screen "SettingPrinter" 800x414, template "Template_Mirai"
   on GenerateScreen: SetTag("screen_titles", 52)
   Button "Button_3" at 256,226 size 80x40; TextOff 'Connect / Pripoj'
      on Release: ResetBit("CON_ConnectHMI")
      on Press: SetBit("CON_ConnectHMI")
   TextField "Text field_3" at 19,231 size 25x32; Text 'IP'
   IOField "I/O field_1" at 61,231 size 180x32; FormatPattern ????????????????????
      ProcessValue <- "PrinterData_CON_PrinterBagData_RemoteAddress"
   TextField "Text field_4" at 167,152 size 42x32; Text 'CON'
   SymbolicIOField "Symbolic I/O field_1" at 65,186 size 170x32; TextOn '1'; TextOff '0'; TextList "CON_Printers"
      ProcessValue <- "PrinterData_CON_PrinterSelection"
   Button "Button_6" at 256,42 size 80x40; TextOff 'Connect / Pripoj'
      on Release: ResetBit("TRP_ConnectHMI")
      on Press: SetBit("TRP_ConnectHMI")
   Button "Button_1" at 256,98 size 120x40; TextOff 'Initialization / Inicializácia'
      on Release: ResetBit("PrinterData_TRP_PrinterData_Initialization")
      on Press: SetBit("PrinterData_TRP_PrinterData_Initialization")
   TextField "Text field_1" at 168,8 size 42x32; Text 'TRP'
   TextField "Text field_2" at 13,47 size 25x32; Text 'IP'
   IOField "I/O field_5" at 38,47 size 213x32; FormatPattern ????????????????????
      ProcessValue <- "PrinterData_TRP_PrinterData_RemoteAddress"
   IOField "I/O field_2" at 61,303 size 180x32; FormatPattern ????????????????????????????????????????????????????????????????????????????????
      ProcessValue <- "PrinterData_CON_PrinterBagData_NonMDR_LabelName"
   TextField "Text field_5" at 19,274 size 223x32; Text 'Non-MDR label name'
   Button "Button_5" at 672,302 size 120x40; TextOff 'Camera settings Nastavenia kamery'
      on Release: ActivateScreen("Setting_DelayTimeM", 0)
   GraphicView "Graphic view_1" at 348,42 size 44x30; Picture "Wbox"
      Visibility <- "TRP_DB_MarkemImaje_ConnectionStatus"
   GraphicView "Graphic view_2" at 346,43 size 45x27; Picture "Cbox"
      Visibility <- "TRP_DB_MarkemImaje_ConnectionStatus"
   GraphicView "Graphic view_3" at 348,229 size 44x30; Picture "Wbox"
      Visibility <- "CON_PrinterConnection"
   GraphicView "Graphic view_4" at 347,231 size 45x27; Picture "Cbox"
      Visibility <- "CON_PrinterConnection"
   Button "Button_4" at 257,301 size 120x40; TextOff 'Initialization / Inicializácia'
      on Release: ResetBit("PrinterData_CON_PrinterBagData_Initialization")
      on Press: SetBit("PrinterData_CON_PrinterBagData_Initialization")
   Switch "Switch_1" at 115,82 size 120x56; TextOn 'DOLE'; CaptionText 'Inverse / Obratena tlac'; TextOff 'HORE'
      on SwitchOff: ResetBit("PrinterData_TRP_PrinterData_Inverse")
      on SwitchOn: SetBit("PrinterData_TRP_PrinterData_Inverse")
      ProcessValue <- "PrinterData_TRP_PrinterData_Inverse"

screen "Setting_DelayTimeM" 800x414, template "Template_Mirai"
   on GenerateScreen: SetTag("screen_titles", 53)
   IOField "I/O field_2" at 160,63 size 104x40; FormatPattern 999
      ProcessValue <- "SP_HMI_Box_Cam_Delay_time_trigger"
   TextField "Text field_2" at 4,63 size 148x40; Text '2D Code Box / 2D kód krabice'
   TextField "Text field_3" at 160,16 size 104x40; Text 'Trigger delay (ms) Oneskorenie čítania (ms)'
   Button "Btn_OpenEditor" at 4,313 size 160x32; TextOff 'Back / Späť'
      on Click: ActivateScreen("SettingPrinter", 0)
   Button "Btn_OpenEditor_1" at 180,313 size 160x32; TextOff 'Camera position / Pozícia kamery'; Authorization "Operate"
      on Click: ActivateScreen("Setting_CameraM", 0)

screen "StatusM" 800x414, template "Template_Mirai"
   on GenerateScreen: SetTag("screen_titles", 51)
   TextField "Text field_2" at 28,39 size 43x23; Text '(01)'
   TextField "Text field_3" at 28,77 size 43x23; Text '(10)'
   TextField "Text field_4" at 28,115 size 43x23; Text '(91)'
   TextField "Text field_5" at 28,153 size 43x23; Text '(92)'
   TextField "Text field_6" at 28,191 size 43x23; Text '(11)'
   TextField "Text field_7" at 28,229 size 43x23; Text '(15)'
   IOField "I/O field_1" at 81,33 size 171x34; FormatPattern ????????????????????????????????????????????????????????????????????????????????
      ProcessValue <- "OPC_TRP_Materia_ActualGTIN_Number"
   IOField "I/O field_2" at 81,71 size 171x34; FormatPattern ????????????????????????????????????????????????????????????????????????????????
      ProcessValue <- "OPC_TRP_Materia_ActualBatchNumber"
   TextField "Text field_8" at 171,9 size 42x23; Text 'TRP'
   IOField "I/O field_3" at 81,109 size 171x34; FormatPattern ????????????????????????????????????????????????????????????????????????????????
      ProcessValue <- "OPC_TRP_Materia_ActualAricleNumber"
   IOField "I/O field_4" at 81,147 size 171x34; FormatPattern ??????
      ProcessValue <- "PrinterData_CON_PrinterBagData_Time"
   IOField "I/O field_5" at 81,185 size 171x34; FormatPattern ????????????????????????????????????????????????????????????????????????????????
      ProcessValue <- "PrinterData_CON_PrinterBagData_Date"
   IOField "I/O field_6" at 81,223 size 171x34; FormatPattern ??????????
      ProcessValue <- "TRP_DB_MarkemImaje_ExtDate"
   TextField "Text field_1" at 548,10 size 110x23; Text 'PLAIN Data'
   TextField "Text field_11" at 400,33 size 90x23; Text 'EAN_TRP / EAN TRP'
   TextField "Text field_13" at 400,63 size 56x23; Text 'Batch'
   TextField "Text field_15" at 400,93 size 100x23; Text 'MachineID'
   TextField "Text field_16" at 400,123 size 90x23; Text 'MDR Flag'
   TextField "Text field_17" at 400,153 size 66x23; Text 'Article'
   TextField "Text field_18" at 400,183 size 99x23; Text 'Batch END'
   TextField "Text field_19" at 400,214 size 92x23; Text 'ART Base'
   TextField "Text field_20" at 400,246 size 87x23; Text 'ART Flag'
   TextField "Text field_21" at 400,278 size 110x23; Text 'Market Reg'
   TextField "Text field_22" at 400,310 size 42x23; Text 'BBD'
   IOField "I/O field_11" at 570,32 size 200x25; FormatPattern ??????????????
      ProcessValue <- "OPC_TRP_Materia_NewGTIN_Number"
   IOField "I/O field_12" at 570,62 size 200x25; FormatPattern ????????????????????????????????????????????????????????????????????????????????
      ProcessValue <- "OPC_CON_Material_NewBatchNumber"
   IOField "I/O field_13" at 570,92 size 200x25; FormatPattern ????????????????????????????????????????????????????????????????????????????????
      ProcessValue <- "OPC_TRP_Materia_NewMachineID"
   IOField "I/O field_14" at 570,122 size 200x25; FormatPattern ????????????????????????????????????????????????????????????????????????????????
      ProcessValue <- "OPC_CON_Material_NewMDR_Flag"
   IOField "I/O field_15" at 570,152 size 200x25; FormatPattern 9999999999
      ProcessValue <- "OPC_TRP_Materia_NewArticleNumber"
   IOField "I/O field_16" at 570,182 size 200x25; FormatPattern ????????????????????????????????????????????????????????????????????????????????
      ProcessValue <- "OPC_CON_Material_NewBatchEndTime"
   IOField "I/O field_17" at 570,213 size 200x25; FormatPattern 9999999999
      ProcessValue <- "OPC_CON_Material_NewArtBaseNumber"
   IOField "I/O field_18" at 570,245 size 200x25; FormatPattern ????????????????????????????????????????????????????????????????????????????????
      ProcessValue <- "OPC_CON_Material_NewArticleFlag"
   IOField "I/O field_19" at 570,277 size 200x25; FormatPattern ?????????????????????
      ProcessValue <- "OPC_CON_Material_NewMarketREG_Code"
   IOField "I/O field_20" at 570,309 size 200x25; FormatPattern ????????????????????????????????????????????????????????????????????????????????
      ProcessValue <- "OPC_CON_Material_NewBBD"
   IOField "I/O field_7" at 55,284 size 115x32; HelpText 'Enter ip+port 10.176.48.110:45'; FormatPattern ??????????
      ProcessValue <- "OPC_TRP_Materia_ActualBatchNumber"
   IOField "I/O field_8" at 194,284 size 115x32; HelpText 'Enter ip+port 10.176.48.110:45'; FormatPattern ??????????
      ProcessValue <- "OPC_CON_Material_ActualArtBaseNumber"
      Visibility <- "CON_DB_HandleComBag_ActualArtFlag"
   IOField "I/O field_10" at 20,302 size 115x32; HelpText 'Enter ip+port 10.176.48.110:45'; FormatPattern ??????????
      ProcessValue <- "OPC_CON_Material_ActualMarketRegCode"
   TextField "Text field_14" at 127,307 size 42x23; Text 'BBD'
      Visibility <- "TRP_DB_MarkemImaje_ExpFlag"
   IOField "I/O field_9" at 165,303 size 76x32; HelpText 'Enter ip+port 10.176.48.110:45'; FormatPattern ??????
      ProcessValue <- "OPC_CON_Material_ActualBBD"
   IOField "I/O field_23" at 296,284 size 76x32; HelpText 'Enter ip+port 10.176.48.110:45'; FormatPattern ?????
      ProcessValue <- "TRP_DB_MarkemImaje_TimePrinted"
      Visibility <- "CON_DB_HandleComBag_ActualArtFlag"
   IOField "I/O field_24" at 159,284 size 76x32; HelpText 'Enter ip+port 10.176.48.110:45'; FormatPattern ??????
      ProcessValue <- "TRP_DB_MarkemImaje_TimePrinted"
      Visibility <- "CON_DB_HandleComBag_ActualArtFlag"
   TextField "Text field_9" at 20,288 size 40x23; Text 'LOT'
   TextField "Text field_12" at 159,288 size 43x23; Text 'ART'
      Visibility <- "CON_DB_HandleComBag_ActualArtFlag"
   TextField "Text field_10" at 151,263 size 43x23; Text 'CON'
   IOField "I/O field_21" at 150,152 size 44x23; HelpText 'Enter ip+port 10.176.48.110:45'; FormatPattern ???
      ProcessValue <- "OPC_TRP_Materia_ActualMachineID"
   IOField "I/O field_22" at 188,152 size 58x23; HelpText 'Enter ip+port 10.176.48.110:45'; FormatPattern 99999
      ProcessValue <- "TRP_DB_MarkemImaje_Serial"

screen "Rec_Edit" 800x414, template "Template_Enigma"
   on GenerateScreen: SetTag("screen_titles", 6)
   IOField "I/O field_1" at 407,54 size 104x32; Authorization "Recipe management"; FormatPattern 9999
      ProcessValue <- "Rec_HMI_Bag_Cam_Vertiacal_position"
   IOField "I/O field_2" at 407,131 size 104x32; Authorization "Recipe management"; FormatPattern s999
      ProcessValue <- "Rec_HMI_Bag_Cam_Angle"
   IOField "I/O field_3" at 407,93 size 104x32; Authorization "Recipe management"; FormatPattern 9999
      ProcessValue <- "Rec_HMI_Bag_Cam_Horizontal_position"
   TextField "Text field_1" at 299,54 size 104x32; Text 'A'
   TextField "Text field_2" at 299,93 size 104x32; Text 'B'
   TextField "Text field_3" at 299,131 size 104x32; Text 'C'
   TextField "Text field_4" at 623,54 size 36x32; Text 'mm'
   TextField "Text field_5" at 623,93 size 36x32; Text 'mm'
   TextField "Text field_6" at 623,131 size 36x32; Text '°'
   TextField "Text field_15" at 299,167 size 104x40; Text 'Trigger delay Oneskorenie čítania'
   IOField "I/O field_4" at 407,171 size 104x32; Authorization "Recipe management"; FormatPattern 999
      ProcessValue <- "Rec_HMI_Bag_Cam_Delay_time_trigger"
   IOField "I/O field_5" at 515,171 size 104x32; Authorization "Recipe management"; FormatPattern 999
      ProcessValue <- "Rec_HMI_Box_Cam_Delay_time_trigger"
   TextField "Text field_16" at 623,171 size 36x32; Text 'ms'
   TextField "Text field_18" at 419,18 size 80x32; Text 'BAG / SÁČOK'
   TextField "Text field_19" at 527,18 size 80x32; Text 'BOX / KRABICA'
   IOField "I/O field_8" at 515,54 size 104x32; Authorization "Recipe management"; FormatPattern 9999
      ProcessValue <- "Rec_HMI_Box_Cam_Vertiacal_position"
   IOField "I/O field_9" at 515,131 size 104x32; Authorization "Recipe management"; FormatPattern s999
      ProcessValue <- "Rec_HMI_Box_Cam_Angle"
   IOField "I/O field_10" at 515,93 size 104x32; Authorization "Recipe management"; FormatPattern 9999
      ProcessValue <- "Rec_HMI_Box_Cam_Horizontal_position"
   Button "Btn_Save" at 692,8 size 80x32; TextOff 'SAVE / ULOŽ'; Authorization "Recipe management"
      on Click: SetTag("Rec_FunctionUsed", 7); "Rec_SafeSave"()
   Button "Btn_ExitEditor" at 8,313 size 216x32; TextOff 'Exit recipe editor / Ukonči editor receptov'
      on Click: ActivateScreen("Rec_Overview", 0)
   GraphicView "Graphic view_1" at 20,77 size 222x229; Picture "CognexDatamanClearedAndSemiTransparent2"
   TextField "Text field_10" at 18,184 size 32x40; Text 'A'
   TextField "Text field_11" at 102,71 size 32x40; Text 'B'
   TextField "Text field_12" at 179,78 size 32x40; Text 'C'
   Button "Btn_ReadSP" at 668,72 size 124x32; TextOff 'READ from PLC / NAČÍTAJ z PLC'; Authorization "Recipe management"
      on Click: SetTag("Rec_FunctionUsed", 8); function_b456aad1(1, "Rec_ReadSPResult")
   TextField "Text field_7" at 8,8 size 264x62; Text 'Recipe name: / Názov receptu: / 配方名'
   IOField "I/O field_6" at 14,35 size 252x30; Authorization "Recipe management"; FormatPattern ????????????????????????????????????????
      ProcessValue <- "Rec_SelectedRecipe"
   GraphicIOField "Graphic I/O field_1" at 408,250 size 32x32; PictureList "On_Off_Editable"
      ProcessValue <- "Rec_HMI_Enigma_off"
   Button "Button_1" at 408,250 size 32x32; TextOff 'Text'
      on Click: InvertBit("Rec_HMI_Enigma_off")
   IOField "I/O field_7" at 407,211 size 104x32; Authorization "Recipe management"; FormatPattern 9999
      ProcessValue <- "Rec_HMI_Bag_Cam_Fps"
   TextField "Text field_13" at 299,211 size 104x32; Text 'Num of pics / Počet snímok'
   IOField "I/O field_11" at 515,211 size 104x32; Authorization "Recipe management"; FormatPattern 9999
      ProcessValue <- "Rec_HMI_Box_Cam_Fps"
   TextField "Text field_14" at 299,250 size 104x32; Text 'Enigma'
   GraphicIOField "Graphic I/O field_2" at 624,250 size 32x32; PictureList "On_Off_Editable"
      ProcessValue <- "Rec_HMI_Mirai_off"
   Button "Button_2" at 624,250 size 32x32; TextOff 'Text'
      on Click: InvertBit("Rec_HMI_Mirai_off")
   TextField "Text field_20" at 515,250 size 104x32; Text 'Mirai'
   Button "Btn_OK_Save_NoNameSpecified" at 692,313 size 80x32; TextOff 'OK / 确定'
      on Click: SetTag("Rec_SaveResult", 0)
      Visibility <- "Rec_SaveResult"
   TextField "Text field_17" at 288,292 size 376x53; Text 'No recipe name set, recipe not saved. Set recipe name and try again. Žiaden zadaný názov receptu, recept sa neuložil. Nastavte názov receptu a skúste to znova. 未设置配方名 不能保存配方。 输入配方名再保存。'
      Visibility <- "Rec_SaveResult"
   TextField "Text field_8" at 288,292 size 376x53; Text 'Saving recipe ... / Ukladanie receptu ... / 配方保存中…'
      Visibility <- "Rec_SaveResult"
   Button "Btn_OK_Save_Success" at 692,313 size 80x32; TextOff 'OK / 确定'
      on Click: SetTag("Rec_SaveResult", 0)
      Visibility <- "Rec_SaveResult"
   TextField "Text field_9" at 288,292 size 376x53; Text 'Recipe saving succeeded. Ukladanie receptu bolo úspešné. 保存配方 成功。'
      Visibility <- "Rec_SaveResult"
   TextField "Text field_24" at 288,292 size 376x53; Text 'Recipe saving failed. Ukladanie receptu zlyhalo. 保存配方 失败。'
      Visibility <- "Rec_SaveResult"
   Button "Btn_OK_Save_Fail" at 692,313 size 80x32; TextOff 'OK / 确定'
      on Click: SetTag("Rec_SaveResult", 0)
      Visibility <- "Rec_SaveResult"
   TextField "Text field_25" at 288,292 size 376x53; Text 'Reading setpoints ... / Čítanie požadovaných hodnôt ... / 读取设定值…'
      Visibility <- "Rec_ReadSPResult"
   Button "Btn_OK_ReadSP_Success" at 692,313 size 80x32; TextOff 'OK / 确定'
      on Click: SetTag("Rec_ReadSPResult", 0)
      Visibility <- "Rec_ReadSPResult"
   TextField "Text field_26" at 288,292 size 376x53; Text 'Reading of setpoints succeeded. Čítanie požadovaných hodnôt bolo úspešné. 读取设定值 成功。'
      Visibility <- "Rec_ReadSPResult"
   TextField "Text field_27" at 288,292 size 376x53; Text 'Reading of setpoints failed. Čítanie požadovaných hodnôt zlyhalo. 读取设定值 失败。'
      Visibility <- "Rec_ReadSPResult"
   Button "Btn_OK_ReadSP_Fail" at 692,313 size 80x32; TextOff 'OK / 确定'
      on Click: SetTag("Rec_ReadSPResult", 0)
      Visibility <- "Rec_ReadSPResult"
   Rectangle "Rectangle_2" at 0,0 size 800x414
      Visibility <- "Rec_FunctionResultSwitch"

screen "Rec_Overview" 800x414, template "Template_Enigma"
   on GenerateScreen: SetTag("screen_titles", 4); SetTag("Rec_FunctionUsed", 0)
   RecipeView "Recipe view_1" at 4,44 size 792x80; DataRecordNameCaption 'Select recipe: / Vyber recept:'; Tag4DataRecord "Rec_SelectedRecipe"; Recipe "ReaderRecipes"
      Visibility <- "Rec_FunctionResultSwitch"
   Button "Btn_Edit" at 88,136 size 76x32; TextOff 'EDIT UPRAV 编辑 所选 配方'; Authorization "Recipe management"
      on Click: SetTag("Rec_FunctionUsed", 5); "Rec_SafeEdit"()
   Button "Btn_Load" at 636,136 size 160x32; TextOff 'LOAD to PLC NAHRAJ do PLC 下载 所选 配方 到PLC'; Authorization "Operate"
      on Click: SetTag("Rec_FunctionUsed", 1); "Rec_SafeLoad"()
   Button "Btn_Delete" at 362,136 size 76x32; TextOff 'DELETE VYMAŽ 删除 所选 配方'; Authorization "Recipe management"
      on Click: SetTag("Rec_FunctionUsed", 2); "Rec_SafeDelete"()
   Button "Btn_View" at 4,136 size 76x32; TextOff 'VIEW ZOBRAZ 浏览 所选 配方'; Authorization "Operate"
      on Click: SetTag("Rec_FunctionUsed", 6); "Rec_SafeView"()
   Button "Btn_OpenEditor" at 4,313 size 216x32; TextOff 'Open recipe editor / Otvor editor receptov'; Authorization "Recipe management"
      on Click: SetTag("Rec_SelectedRecipe", ''); ActivateScreen("Rec_Edit", 0)
   TextField "Text field_12" at 8,8 size 201x32; Text 'Article number: / Číslo artiklu:'
   IOField "I/O field_6" at 200,8 size 162x32; FormatPattern ??????????
      ProcessValue <- "PlainHandle_DB_NewArticleNum"
   Button "Btn_OK_Edit_NoRecipeSelected" at 362,176 size 76x32; TextOff 'OK / 确定'
      on Click: SetTag("Rec_EditResult", 0)
      Visibility <- "Rec_EditResult"
   Button "Btn_OK_Delete_NoRecipeSelected" at 362,176 size 76x32; TextOff 'OK / 确定'
      on Click: SetTag("Rec_DeleteResult", 0)
      Visibility <- "Rec_DeleteResult"
   Button "Btn_OK_View_NoRecipeSelected" at 362,176 size 76x32; TextOff 'OK / 确定'
      on Click: SetTag("Rec_ViewResult", 0)
      Visibility <- "Rec_ViewResult"
   Button "Btn_OK_Load_NoRecipeSelected" at 362,176 size 76x32; TextOff 'OK / 确定'
      on Click: SetTag("Rec_LoadResult", 0)
      Visibility <- "Rec_LoadResult"
   TextField "Text field_15" at 4,44 size 792x124; Text 'No recipe selected. / Nie je vybratý žiaden recept. / 未选配方。'
      Visibility <- "Rec_FunctionResultSwitch"
   TextField "Text field_11" at 4,44 size 792x124; Text 'Recipe loading failed. / Načítavanie receptu zlyhalo. / 下载配方失败。'
      Visibility <- "Rec_LoadResult"
   Button "Btn_OK_Load_Fail" at 362,176 size 76x32; TextOff 'OK / 确定'
      on Click: SetTag("Rec_LoadResult", 0)
      Visibility <- "Rec_LoadResult"
   TextField "Text field_7" at 4,44 size 792x124; Text 'Recipe deletion failed. / Mazanie receptu zlyhalo. / 删除配方失败。'
      Visibility <- "Rec_DeleteResult"
   Button "Btn_OK_Delete_Fail" at 362,176 size 76x32; TextOff 'OK / 确定'
      on Click: SetTag("Rec_DeleteResult", 0)
      Visibility <- "Rec_DeleteResult"
   Rectangle "Rectangle_1" at 0,0 size 800x414
      Visibility <- "Rec_FunctionResultSwitch"
   TextField "Text field_4" at 4,44 size 792x124; Text 'Recipe loading ... / Načítavanie receptu... / 配方表下载中…'
      Visibility <- "Rec_LoadResult"
   Button "Btn_OK_Load_Success" at 362,176 size 76x32; TextOff 'OK / 确定'
      on Click: SetBit("HMI_Control_NewRecipeLoaded"); SetTag("Rec_LoadResult", 0)
      Visibility <- "Rec_LoadResult"
   TextField "Text field_3" at 4,44 size 792x124; Text 'Recipe loading succeeded. / Načítavanie receptu bolo úspešné. / 下载配方成功。'
      Visibility <- "Rec_LoadResult"
   TextField "Text field_5" at 4,44 size 792x124; Text 'Deleting recipe ... / Vymazávanie receptu... / 删除配方…'
      Visibility <- "Rec_DeleteResult"
   Button "Btn_OK_Delete_Success" at 362,176 size 76x32; TextOff 'OK / 确定'
      on Click: SetTag("Rec_SelectedRecipe", ''); SetTag("Rec_DeleteResult", 0)
      Visibility <- "Rec_DeleteResult"
   TextField "Text field_6" at 4,44 size 792x124; Text 'Recipe deletion succeeded. / Mazanie receptu bolo úspešné. / 删除配方成功。'
      Visibility <- "Rec_DeleteResult"
   TextField "Text field_16" at 4,44 size 792x124; Text 'Opening recipe for editing ... / Prebieha otváranie receptu na úpravu ... / 打开编辑配方…'
      Visibility <- "Rec_EditResult"
   Button "Btn_OK_Edit_Success" at 362,176 size 76x32; TextOff 'OK / 确定'
      on Click: SetTag("Rec_EditResult", 0); ActivateScreen("Rec_Edit", 2)
      Visibility <- "Rec_EditResult"
   TextField "Text field_17" at 4,44 size 792x124; Text 'Recipe opening for editing succeeded. / Otváranie receptu na úpravu bolo úspešné. / 打开编辑配方成功。'
      Visibility <- "Rec_EditResult"
   TextField "Text field_1" at 4,44 size 792x124; Text 'Recipe opening for editing failed. / Otváranie receptu na úpravu zlyhalo. / 打开编辑配方失败。'
      Visibility <- "Rec_EditResult"
   Button "Btn_OK_Edit_Fail" at 362,176 size 76x32; TextOff 'OK / 确定'
      on Click: SetTag("Rec_EditResult", 0)
      Visibility <- "Rec_EditResult"
   TextField "Text field_2" at 4,44 size 792x124; Text 'Opening recipe for viewing ... / Prebieha otváranie receptu na prezeranie ... / 打开查看配方…'
      Visibility <- "Rec_ViewResult"
   Button "Btn_OK_View_Success" at 362,176 size 76x32; TextOff 'OK / 确定'
      on Click: SetTag("Rec_ViewResult", 0); ActivateScreen("Rec_View", 2)
      Visibility <- "Rec_ViewResult"
   TextField "Text field_20" at 4,44 size 792x124; Text 'Recipe opening for viewing succeeded. / Otváranie receptu na prezeranie bolo úspešné. / 打开查看配方成功。'
      Visibility <- "Rec_ViewResult"
   TextField "Text field_21" at 4,44 size 792x124; Text 'Recipe opening for viewing failed. / Otváranie receptu na prezeranie zlyhalo. / 打开查看配方失败。'
      Visibility <- "Rec_ViewResult"
   Button "Btn_OK_View_Fail" at 362,176 size 76x32; TextOff 'OK / 确定'
      on Click: SetTag("Rec_ViewResult", 0)
      Visibility <- "Rec_ViewResult"

screen "Rec_View" 800x414, template "Template_Enigma"
   on GenerateScreen: SetTag("screen_titles", 5)
   IOField "I/O field_1" at 407,54 size 104x32; FormatPattern 9999
      ProcessValue <- "Rec_HMI_Bag_Cam_Vertiacal_position"
   IOField "I/O field_2" at 407,131 size 104x32; FormatPattern s999
      ProcessValue <- "Rec_HMI_Bag_Cam_Angle"
   IOField "I/O field_3" at 407,93 size 104x32; FormatPattern 9999
      ProcessValue <- "Rec_HMI_Bag_Cam_Horizontal_position"
   TextField "Text field_1" at 299,54 size 104x32; Text 'A'
   TextField "Text field_2" at 299,93 size 104x32; Text 'B'
   TextField "Text field_3" at 299,131 size 104x32; Text 'C'
   TextField "Text field_4" at 623,54 size 36x32; Text 'mm'
   TextField "Text field_5" at 623,93 size 36x32; Text 'mm'
   TextField "Text field_6" at 623,131 size 36x32; Text '°'
   TextField "Text field_15" at 299,167 size 104x40; Text 'Trigger delay Oneskorenie čítania'
   IOField "I/O field_4" at 407,171 size 104x32; FormatPattern 999
      ProcessValue <- "Rec_HMI_Bag_Cam_Delay_time_trigger"
   IOField "I/O field_5" at 515,171 size 104x32; FormatPattern 999
      ProcessValue <- "Rec_HMI_Box_Cam_Delay_time_trigger"
   TextField "Text field_16" at 623,171 size 36x32; Text 'ms'
   TextField "Text field_18" at 419,18 size 80x32; Text 'BAG / SÁČOK'
   TextField "Text field_19" at 523,18 size 80x32; Text 'BOX / KRABICA'
   IOField "I/O field_8" at 515,54 size 104x32; FormatPattern 9999
      ProcessValue <- "Rec_HMI_Box_Cam_Vertiacal_position"
   IOField "I/O field_9" at 515,131 size 104x32; FormatPattern s999
      ProcessValue <- "Rec_HMI_Box_Cam_Angle"
   IOField "I/O field_10" at 515,93 size 104x32; FormatPattern 9999
      ProcessValue <- "Rec_HMI_Box_Cam_Horizontal_position"
   Button "Button_7" at 8,313 size 216x32; TextOff 'Exit recipe viewer / Ukonči prehliadač receptov'
      on Click: ActivateScreen("Rec_Overview", 0)
   GraphicView "Graphic view_1" at 20,77 size 222x229; Picture "CognexDatamanClearedAndSemiTransparent2"
   TextField "Text field_10" at 18,184 size 32x40; Text 'A'
   TextField "Text field_11" at 102,71 size 32x40; Text 'B'
   TextField "Text field_12" at 179,78 size 32x40; Text 'C'
   TextField "Text field_7" at 8,8 size 264x62; Text 'Recipe name: / Názov receptu: / 配方名'
   IOField "I/O field_6" at 14,35 size 252x30; FormatPattern ????????????????????????????????????????
      ProcessValue <- "Rec_SelectedRecipe"
   GraphicIOField "Graphic I/O field_1" at 408,250 size 32x32; PictureList "On_Off_NonEditable"
      ProcessValue <- "Rec_HMI_Enigma_off"
   IOField "I/O field_7" at 407,211 size 104x32; Authorization "Recipe management"; FormatPattern 9999
      ProcessValue <- "Rec_HMI_Bag_Cam_Fps"
   TextField "Text field_13" at 299,211 size 104x32; Text 'Num of pics / Počet snímok'
   IOField "I/O field_11" at 515,211 size 104x32; Authorization "Recipe management"; FormatPattern 9999
      ProcessValue <- "Rec_HMI_Box_Cam_Fps"
   TextField "Text field_14" at 299,250 size 104x32; Text 'Enigma'
   GraphicIOField "Graphic I/O field_2" at 624,250 size 32x32; PictureList "On_Off_NonEditable"
      ProcessValue <- "Rec_HMI_Mirai_off"
   TextField "Text field_20" at 515,250 size 104x32; Text 'Mirai'

screen "SystemScreenE" 800x414, template "Template_Enigma"
   on GenerateScreen: SetTag("screen_titles", 20)
   Button "HmiScreenItemData_2" at 196,73 size 169x52; TextOn 'Projektinformationen / Project information / Informatii proiect / ข้อมูลโปรเจ็ค / Informácie o projekte'; TextOff 'Projektinformationen Project information Informatii proiect ข้อมูลโปรเจ็ค Informácie o projekte'; PictureOn "Navigates to Projektinformationen for HMI_1"; PictureOff "Graphic_1"
      on Press: ActivateScreen("ProjectInfo", 0)
   Button "HmiScreenItemData_3" at 435,201 size 169x52; TextOn 'Systemeinstellungen System settings Setarile de sistem Configurações de sistema ตั้งค่าระบบ Systémové nastavenia'; TextOff 'Systemeinstellungen System settings Setarile de sistem Configurações de sistema ตั้งค่าระบบ Systémové nastavenia'; Authorization "User administration"; PictureOff "Graphic_6"; PictureOn "Graphic_6"
      on Press: ActivateScreen("SystemSettings", 0)
   Button "HmiScreenItemData_4" at 196,137 size 169x52; TextOn 'Benutzerverwaltung User administration De administrare a utilizatorilor Administração de usuários การควบคุมผู้ใช้งาน Správa používateľov'; TextOff 'Benutzerverwaltung User administration De administrare a utilizatorilor Administração de usuários การควบคุมผู้ใช้งาน Správa používateľov'; Authorization "User administration"; PictureOff "Graphic_4"; PictureOn "Navigates to Benutzerverwaltung for HMI_1"
      on Press: ActivateScreen("UserAdmin", 0)
   Button "HmiScreenItemData_5" at 435,73 size 169x52; TextOn 'Systeminformationen / System information / Informatii sistem / Informação do sistema / ข้อมูลระบบ / Informácie o systéme'; TextOff 'Systeminformationen System information Informatii sistem Informação do sistema ข้อมูลระบบ Informácie o systéme'; PictureOn "Graphic_2"; PictureOff "Graphic_2"
      on Press: ActivateScreen("SystemInfo", 0)
   Button "HmiScreenItemData_6" at 435,137 size 169x52; TextOn 'Verschiedene Aufgaben Other tools Diverse activitati Various tasks งานอื่นๆ Iné nástroje'; TextOff 'Verschiedene Aufgaben Other tools Diverse activitati Various tasks งานอื่นๆ Iné nástroje'; PictureOn "Navigates to Verschiedene Aufgaben for HMI_1"; PictureOff "Graphic_5"
      on Press: ActivateScreen("OtherTools", 0)
   Button "HmiScreenItemData_1" at 195,201 size 169x52; TextOn 'Systemeinstellungen System diagnostics Setarile de sistem Configurações de sistema ตั้งค่าระบบ Diagnostika systému'; TextOff 'Systemeinstellungen System diagnostics Setarile de sistem Configurações de sistema ตั้งค่าระบบ Diagnostika systému'; PictureOff "Graphic_3"; PictureOn "Graphic_3"; Authorization "Operate"
      on Press: ActivateScreen("Diagnostic", 0)

screen "ProjectInfo" 800x414
   on GenerateScreen: SetTag("screen_titles", 21)
   TextField "HmiScreenItemData" at 140,89 size 250x27; Text 'Projektname: / Project name: / Nome do projeto: / ชื่อโปรเจ็ค: / Názov projektu:'
   TextField "HmiScreenItemData_1" at 410,89 size 312x27; Text 'Yokohama_Skiver / ENIGMA_Essity_TP700 / TP1200_MRH / MRH_ประเทศไทย_TP700'
   TextField "HmiScreenItemData_2" at 140,119 size 250x27; Text 'Erstellt: / Created: / Criado: / การผลิต: / Vytvoril:'
   TextField "HmiScreenItemData_3" at 410,119 size 312x27; Text '07.03.2014 09:50:27 / 2019 / 2016 / 2018'
   TextField "HmiScreenItemData_4" at 140,148 size 250x27; Text 'Autor: / Author: / ผู้เขียน:'
   TextField "HmiScreenItemData_5" at 410,148 size 312x27; Text 'admin / Ing. Andrea Bečárová / Veronika Wolfová / Maria Ivankova / Lukas Vilasek'
   TextField "HmiScreenItemData_6" at 140,178 size 250x27; Text 'Beschreibung: / Description: / Descrição: / การอธิบายลักษณะ: / Popis:'
   TextField "HmiScreenItemData_7" at 410,178 size 312x27; Text '(nicht konfiguriert) / (not configured) / (ยังไม่ได้ทำการตั้งค่า)'
   Button "Button_7" at 8,313 size 152x32; TextOff 'Back / Späť'
      on Click: function_efd93a16()

screen "SystemInfo" 800x414
   on GenerateScreen: SetTag("screen_titles", 22)
   TextField "HmiScreenItemData" at 140,89 size 250x27; Text 'Bediengerätetyp: / Device type: / Tipo de dispositivo: / Typ zariadenia: / ประเภทของดีไวซ์:'
   TextField "HmiScreenItemData_1" at 410,89 size 250x27; Text 'TP900 Comfort 12.0 / TP700 Comfort 15.1.0.0 / TP1200 Comfort 13.0 / TP700 คอมฟอร์ท 14.0.1.0'
   TextField "HmiScreenItemData_2" at 140,119 size 250x27; Text 'Version: / Verzia: / เวอร์ชั่น'
   TextField "HmiScreenItemData_3" at 140,148 size 250x27; Text 'Verbindung: / Connection: / Conexão: / Komunikácia: / การเชื่อมต่อ:'
   TextField "HmiScreenItemData_4" at 410,148 size 250x27; Text '(nicht konfiguriert) / (not configured) / (ยังไม่ได้ทำการตั้งค่า)'
   TextField "HmiScreenItemData_5" at 140,178 size 250x27; Text 'Steuerung: / Control system: / Sistema de controle: / Riadiaci systém: / ระบบควบคุม:'
   TextField "HmiScreenItemData_6" at 410,178 size 250x27; Text '<PLC>'
   Button "HmiScreenItemData_7" at 410,119 size 250x27; TextOn 'Version anzeigen'; TextOff 'Version anzeigen / Show version / Mostrar a versão / Zobraziť verziu / เวอร์ชั่นที่แสดง'
      on Press: function_febcb963(-1)
   Button "Button_7" at 8,313 size 152x32; TextOff 'Back / Späť'
      on Click: function_efd93a16()

screen "SystemSettings" 800x414
   on GenerateScreen: SetTag("screen_titles", 26)
   Button "HmiScreenItemData" at 225,54 size 169x52; TextOn 'Online'; TextOff 'Online / ออฟไลน์'
      on Press: function_bb44b551(0)
   Button "HmiScreenItemData_1" at 225,118 size 169x52; TextOn 'Offline'; TextOff 'Offline / ออฟไลน์'
      on Press: function_bb44b551(1)
   Button "HmiScreenItemData_2" at 225,182 size 169x52; TextOn 'Transfer'; TextOff 'Transfer / Transferir / Prenos / การเปลี่ยนถ่าย'
      on Press: function_bb44b551(2)
   Button "HmiScreenItemData_4" at 406,54 size 169x52; TextOn 'Systemsteuerung'; TextOff 'Systemsteuerung / Control panel / Painel de controle / Ovládací panel / แผงควบคุม'
      on Press: function_f34a74f3()
   Button "Button_7" at 8,313 size 152x32; TextOff 'Back / Späť'
      on Click: function_efd93a16()

screen "OtherTools" 800x414
   on GenerateScreen: SetTag("screen_titles", 24)
   Button "HmiScreenItemData" at 241,54 size 169x52; TextOn 'Bildschirm kalibrieren'; TextOff 'Bildschirm kalibrieren / Calibrate touchscreen / Calibrar tela de toque / คาลิเบรต หน้าจอสัมผัส / Kalibrácia obrazovky'; Authorization "User administration"
      on Press: function_bc3e350c()
   Button "HmiScreenItemData_1" at 241,118 size 169x52; TextOn 'Putzbild'; TextOff 'Putzbild / Clean screen / Tela limpa / ทำความสะอาดสกรีน / Čistenie obrazovky'
      on Press: function_be740847(15)
   Button "Button_3" at 467,118 size 80x52; TextOff 'ExitRuntime Exit runtime Exitruntime ( เอ็กซิส รันไทม์) Ukonči runtime'; PictureOn "ExitRuntime_TP900_Comfort"; PictureOff "ExitRuntime_TP900_Comfort"; Authorization "User administration"
      on Press: StopRuntime(0)
   Button "Button_2" at 467,54 size 80x52; TextOn 'Login / ลงชื่อเข้าใช้'; TextOff 'Login / ลงชื่อเข้าใช้'; PictureOn "Login_TP900_Comfort"; PictureOff "Login_TP900_Comfort"
      on Press: function_a2a04561()
   Button "Button_7" at 8,313 size 152x32; TextOff 'Back / Späť'
      on Click: function_efd93a16()

screen "UserAdmin" 800x414
   on GenerateScreen: SetTag("screen_titles", 23)
   UserView "HmiScreenItemData" at 4,4 size 792x300
   Button "Button_7" at 8,313 size 152x32; TextOff 'Back / Späť'
      on Click: function_efd93a16()

screen "Diagnostic" 800x414
   on GenerateScreen: SetTag("screen_titles", 25)
   SysDiagControl "System diagnostics view_1" at 4,4 size 792x300
   Button "Button_7" at 8,313 size 152x32; TextOff 'Back / Späť'
      on Click: function_efd93a16()

screen "MainScreen" 800x414, template "Template_Enigma"
   on GenerateScreen: SetTag("screen_titles", 1); SetTag("autoPwd", 'operator'); SetTag("autoUser", 'operator'); "AutoLoginOperator"()
   TextField "Text field_1" at 412,8 size 148x23; Text '2D code on BOX / 2D kód na krabici'
   TextField "Text field_2" at 412,80 size 200x23; Text 'Actual reading box / Prečítaný kód krabice'
   TextField "Text field_3" at 412,104 size 200x23; Text 'Materialnumber box / Aktuálny kód krabice'
   TextField "Text field_4" at 412,200 size 200x23; Text '#Triggers box / #Senzor krabica'
   TextField "Text field_5" at 412,224 size 200x23; Text '#NoRead box / #Neprečítaná krabica'
   TextField "Text field_6" at 412,248 size 200x23; Text '#Mismatch box / #Nezhodná krabica'
   TextField "Text field_7" at 12,8 size 148x23; Text '2D code on BAG / 2D kód na sáčku'
   TextField "Text field_8" at 12,80 size 200x23; Text 'Actual reading bag / Prečítaný kód sáčku'
   TextField "Text field_9" at 12,104 size 200x23; Text 'Material number bag / Aktuálny kód sáčku'
   TextField "Text field_10" at 12,200 size 200x23; Text '#Triggers bag / #Senzor sáčok'
   TextField "Text field_11" at 12,224 size 200x23; Text '#NoRead bag / #Neprečítaný sáčok'
   TextField "Text field_12" at 12,248 size 200x23; Text '#Mismatch bag / #Nezhodný sáčok'
   IOField "I/O field_1" at 632,80 size 148x23; FormatPattern 9999999999
      ProcessValue <- "HMI_Box_Small_Codes_ActualReadingBox"
   IOField "I/O field_2" at 632,104 size 148x23; FormatPattern 9999999999
      ProcessValue <- "HMI_Box_Small_Codes_MaterialNumberBox"
   IOField "I/O field_3" at 632,200 size 148x23; FormatPattern 9999999999
      ProcessValue <- "HMI_Box_Small_Counters_Trigger"
   IOField "I/O field_4" at 632,224 size 148x23; FormatPattern 9999999999
      ProcessValue <- "HMI_Box_Small_Counters_CodeBadRead"
   IOField "I/O field_5" at 632,248 size 148x23; FormatPattern 9999999999
      ProcessValue <- "HMI_Box_Small_Counters_CodeNok"
   IOField "I/O field_6" at 232,80 size 148x23; FormatPattern 9999999999
      ProcessValue <- "HMI_Bag_Codes_ActualReadingBox"
   IOField "I/O field_7" at 232,104 size 148x23; FormatPattern 9999999999
      ProcessValue <- "HMI_Bag_Codes_MaterialNumberBox"
   IOField "I/O field_8" at 232,200 size 148x23; FormatPattern 9999999999
      ProcessValue <- "HMI_Bag_Counters_Trigger"
   IOField "I/O field_9" at 232,224 size 148x23; FormatPattern 9999999999
      ProcessValue <- "HMI_Bag_Counters_CodeBadRead"
   IOField "I/O field_10" at 232,248 size 148x23; FormatPattern 9999999999
      ProcessValue <- "HMI_Bag_Counters_CodeNok"
   TextField "Text field_13" at 412,48 size 200x23; Text 'TCP communication / TCP komunikácia'
   TextField "Text field_14" at 12,48 size 200x23; Text 'TCP communication / TCP komunikácia'
   SymbolicIOField "Symbolic I/O field_1" at 632,49 size 148x23; TextOn 'OK / NOK'; TextOff 'NOK / OK'
      ProcessValue <- "HMI_Box_Small_Control_TcpCom"
      Appearance <- "HMI_Box_Small_Control_TcpCom"
   SymbolicIOField "Symbolic I/O field_2" at 232,48 size 148x23; TextOn 'OK / NOK'; TextOff 'NOK / OK'
      ProcessValue <- "HMI_Bag_Control_TcpCom"
      Appearance <- "HMI_Bag_Control_TcpCom"

screen "Alarm history_Enigma" 800x414, template "Template_Enigma"
   on GenerateScreen: SetTag("screen_titles", 2)
   AlarmView "Alarm view_1" at 0,0 size 800x349

screen "Setting_Camera" 800x414, template "Template_Enigma"
   on GenerateScreen: SetTag("screen_titles", 8)
   IOField "I/O field_1" at 407,126 size 104x32; FormatPattern 9999
      ProcessValue <- "SP_HMI_Bag_Cam_Vertiacal_position"
   IOField "I/O field_2" at 407,202 size 104x32; FormatPattern s999
      ProcessValue <- "SP_HMI_Bag_Cam_Angle"
   IOField "I/O field_3" at 407,164 size 104x32; FormatPattern 9999
      ProcessValue <- "SP_HMI_Bag_Cam_Horizontal_position"
   TextField "Text field_1" at 299,126 size 104x32; Text 'A'
   TextField "Text field_2" at 299,164 size 104x32; Text 'B'
   TextField "Text field_3" at 299,202 size 104x32; Text 'C'
   TextField "Text field_4" at 623,126 size 36x32; Text 'mm'
   TextField "Text field_5" at 623,164 size 36x32; Text 'mm'
   TextField "Text field_6" at 623,202 size 36x32; Text '°'
   TextField "Text field_18" at 419,90 size 80x32; Text 'BAG / SÁČOK'
   TextField "Text field_19" at 523,90 size 80x32; Text 'BOX / KRABICA'
   IOField "I/O field_8" at 515,126 size 104x32; FormatPattern 9999
      ProcessValue <- "SP_HMI_Box_Cam_Vertiacal_position"
   IOField "I/O field_9" at 515,202 size 104x32; FormatPattern s999
      ProcessValue <- "SP_HMI_Box_Cam_Angle"
   IOField "I/O field_10" at 515,164 size 104x32; FormatPattern 9999
      ProcessValue <- "SP_HMI_Box_Cam_Horizontal_position"
   Button "Button_7" at 8,313 size 152x32; TextOff 'Back / Späť'
      on Click: ActivateScreen("Setting_DelayTime", 0)
   GraphicView "Graphic view_1" at 20,53 size 224x212; Picture "CognexDatamanEdited_3"
   TextField "Text field_10" at 18,144 size 32x40; Text 'A'
   TextField "Text field_11" at 102,31 size 32x40; Text 'B'
   TextField "Text field_12" at 179,38 size 32x40; Text 'C'
   TextField "Text field_7" at 288,8 size 376x62; Text 'Camera position: / Pozícia kamery: / 配方名'
   GraphicIOField "Graphic I/O field_1" at 408,243 size 32x32; PictureList "On_Off_NonEditable"
      ProcessValue <- "SP_HMI_Enigma_off"
   TextField "Text field_14" at 299,243 size 104x32; Text 'Enigma'
   GraphicIOField "Graphic I/O field_2" at 624,243 size 32x32; PictureList "On_Off_NonEditable"
      ProcessValue <- "SP_HMI_Mirai_off"
   TextField "Text field_20" at 515,243 size 104x32; Text 'Mirai'

screen "Setting_DelayTime" 800x414, template "Template_Enigma"
   on GenerateScreen: SetTag("screen_titles", 7)
   TextField "Text field_1" at 4,63 size 148x40; Text '2D Code Bag / 2D kód sáčku'
   TextField "Text field_2" at 4,111 size 148x40; Text '2D Code Box / 2D kód krabice'
   TextField "Text field_3" at 160,16 size 104x40; Text 'Trigger delay (ms) Oneskorenie čítania (ms)'
   IOField "I/O field_1" at 160,63 size 104x40; FormatPattern 999
      ProcessValue <- "SP_HMI_Bag_Cam_Delay_time_trigger"
   IOField "I/O field_2" at 160,111 size 104x40; FormatPattern 999
      ProcessValue <- "SP_HMI_Box_Cam_Delay_time_trigger"
   Button "Btn_OpenEditor" at 4,313 size 160x32; TextOff 'Camera position / Pozícia kamery'; Authorization "Operate"
      on Click: ActivateScreen("Setting_Camera", 0)

screen "StatusE" 800x414, template "Template_Enigma"
   on GenerateScreen: SetTag("screen_titles", 3)
   TextField "Text field_1" at 448,16 size 100x40; Text 'Counters BAG Počítadlá sáčkov'
   TextField "Text field_2" at 624,16 size 100x40; Text 'Counters BOX Počítadlá krabíc'
   TextField "Text field_3" at 7,20 size 160x40; Text 'Actual production / Aktuálna výroba'
   TextField "Text field_8" at 12,80 size 160x23; Text 'Line number / Číslo linky'
   TextField "Text field_9" at 12,112 size 160x23; Text 'Order number / Číslo objednávky'
   IOField "I/O field_6" at 184,80 size 148x23; FormatPattern ??????????
      ProcessValue <- "HMI_line_number_s"
   IOField "I/O field_7" at 184,112 size 148x23; FormatPattern ?????????????
      ProcessValue <- "HMI_order_number_s"
   TextField "Text field_4" at 12,144 size 160x23; Text 'Article number / Číslo artiklu'
   IOField "I/O field_1" at 184,144 size 148x23; FormatPattern ?????????????
      ProcessValue <- "HMI_article_number_s"
   IOField "I/O field_2" at 184,176 size 148x23; FormatPattern ??????????
      ProcessValue <- "HMI_product_weight_s"
   TextField "Text field_5" at 12,176 size 160x23; Text 'Product weight / Hmotnosť produktu'
   IOField "I/O field_3" at 184,208 size 148x23; FormatPattern ??????????
      ProcessValue <- "HMI_total_in_bag_s"
   TextField "Text field_6" at 12,208 size 160x23; Text 'Total in bag / Počet v sáčku'
   IOField "I/O field_4" at 184,240 size 148x23; FormatPattern ??????????
      ProcessValue <- "HMI_total_in_box_s"
   TextField "Text field_7" at 12,240 size 160x23; Text 'Total in box / Počet v krabici'
   TextField "Text field_10" at 372,80 size 72x23; Text 'OK'
   TextField "Text field_11" at 372,120 size 72x23; Text 'NOK'
   TextField "Text field_12" at 372,160 size 72x23; Text 'NO READ'
   TextField "Text field_13" at 372,200 size 72x23; Text 'NDR'
   TextField "Text field_14" at 372,240 size 72x23; Text 'TRIGGER / SENZOR'
   IOField "I/O field_5" at 461,76 size 104x32; FormatPattern 99999
      ProcessValue <- "HMI_Bag_Counters_CodeOk"
   IOField "I/O field_8" at 461,116 size 104x32; FormatPattern 99999
      ProcessValue <- "HMI_Bag_Counters_CodeNok"
   IOField "I/O field_9" at 461,156 size 104x32; FormatPattern 99999
      ProcessValue <- "HMI_Bag_Counters_CodeBadRead"
   IOField "I/O field_10" at 461,196 size 104x32; FormatPattern 99999
      ProcessValue <- "HMI_Bag_Counters_NDR"
   IOField "I/O field_11" at 461,236 size 104x32; FormatPattern 99999
      ProcessValue <- "HMI_Bag_Counters_Trigger"
   Button "Button_2" at 461,281 size 104x32; TextOff 'RESET'
      on Release: ResetBit("HMI_Bag_Control_ResetCounters")
      on Press: SetBit("HMI_Bag_Control_ResetCounters")
   IOField "I/O field_12" at 637,76 size 104x32; FormatPattern 99999
      ProcessValue <- "HMI_Box_Small_Counters_CodeOk"
   IOField "I/O field_13" at 637,116 size 104x32; FormatPattern 99999
      ProcessValue <- "HMI_Box_Small_Counters_CodeNok"
   IOField "I/O field_14" at 637,156 size 104x32; FormatPattern 99999
      ProcessValue <- "HMI_Box_Small_Counters_CodeBadRead"
   IOField "I/O field_15" at 637,196 size 104x32; FormatPattern 99999
      ProcessValue <- "HMI_Box_Small_Counters_NDR"
   IOField "I/O field_16" at 637,236 size 104x32; FormatPattern 99999
      ProcessValue <- "HMI_Box_Small_Counters_Trigger"
   Button "Button_1" at 637,281 size 104x32; TextOff 'RESET'
      on Release: ResetBit("HMI_Box_Small_Control_ResetCounters")
      on Press: SetBit("HMI_Box_Small_Control_ResetCounters")

screen "Service" 800x414
   on GenerateScreen: SetTag("screen_titles", 60)
   IOField "I/O field_1" at 96,56 size 184x32; Authorization "User administration"; FormatPattern ??????????
      ProcessValue <- "X_Simulacia_DB_BagServis"
   IOField "I/O field_2" at 96,96 size 184x32; Authorization "User administration"; FormatPattern ??????????
      ProcessValue <- "X_Simulacia_DB_BoxServis"
   IOField "I/O field_3" at 510,56 size 184x32; Authorization "User administration"; FormatPattern ??????????????
      ProcessValue <- "X_Simulacia_DB_TRP_Materia_NewGTIN_Number"
   Button "Btn_Save" at 700,216 size 80x32; TextOff 'SET / NASTAV'; Authorization "User administration"
      on Release: ResetBit("X_Simulacia_DB_Servis_BoxLarge")
      on Press: SetBit("X_Simulacia_DB_Servis_BoxLarge")
   TextField "Text field_1" at 8,11 size 388x23; Text 'ENIGMA'
   TextField "Text field_2" at 404,11 size 388x23; Text 'MIRAI'
   TextField "Text field_3" at 12,56 size 84x32; Text 'BAG / SÁČOK'
   TextField "Text field_4" at 12,96 size 84x32; Text 'BOX / KRABICA'
   Button "Btn_Save_1" at 302,56 size 80x32; TextOff 'SET / NASTAV'; Authorization "User administration"
      on Release: ResetBit("X_Simulacia_DB_Servis_Bag")
      on Press: SetBit("X_Simulacia_DB_Servis_Bag")
   Button "Btn_Save_2" at 302,96 size 80x32; TextOff 'SET / NASTAV'; Authorization "User administration"
      on Release: ResetBit("X_Simulacia_DB_Servis_BoxSmall")
      on Press: SetBit("X_Simulacia_DB_Servis_BoxSmall")
   Button "Button_7" at 8,313 size 152x32; TextOff 'Back / Späť'
      on Click: ActivateScreen("Menu", 0)
   IOField "I/O field_4" at 510,96 size 184x32; Authorization "User administration"; FormatPattern ??????????
      ProcessValue <- "X_Simulacia_DB_TRP_Materia_NewBatchNumber"
   IOField "I/O field_5" at 510,136 size 184x32; Authorization "User administration"; FormatPattern 9999999999
      ProcessValue <- "X_Simulacia_DB_TRP_Materia_NewArticleNumber"
   IOField "I/O field_6" at 510,176 size 184x32; Authorization "User administration"; FormatPattern ??????????????
      ProcessValue <- "X_Simulacia_DB_TRP_Materia_NewMachineID"
   IOField "I/O field_7" at 510,216 size 184x32; Authorization "User administration"; FormatPattern ??????
      ProcessValue <- "X_Simulacia_DB_TRP_Materia_NewBBD"
   TextField "Text field_5" at 408,56 size 96x32; Text 'GTIN no. / Č. GTIN'
   TextField "Text field_6" at 408,96 size 96x32; Text 'Batch no. / Č. dávky'
   TextField "Text field_7" at 408,136 size 96x32; Text 'Article no. / Č. artiklu'
   TextField "Text field_8" at 408,176 size 96x32; Text 'Machine ID / ID stroja'
   TextField "Text field_9" at 408,216 size 96x32; Text 'Ext. date / Ext. dátum'
   Button "Button_1" at 19,206 size 132x35; TextOff 'Enigma On/Off'; Authorization "User administration"
      on Press: InvertBit("SP_HMI_Enigma_off")
      Appearance <- "SP_HMI_Enigma_off"
   Button "Button_2" at 19,248 size 132x35; TextOff 'Mirai On/Off'; Authorization "User administration"
      on Press: InvertBit("SP_HMI_Mirai_off")
      Appearance <- "SP_HMI_Mirai_off"

Template "Template_Enigma" 800x414
   Button "Exit" at 721,354 size 78x58; TextOff 'Exit'; Authorization "User administration"; PictureOff "ExitRuntime_TP700_Comfort_TR"; PictureOn "ExitRuntime_TP700_Comfort_TR"
      on Release: StopRuntime(0)
   Button "Template_Button" at 321,354 size 78x58; TextOff 'Recipes Správa receptov'
      on Release: ActivateScreen("Rec_Overview", 0)
   Button "Template_Button_1" at 561,354 size 78x58; TextOff 'System / Systém'
      on Release: ActivateScreen("SystemScreenE", 0)
   Button "Template_Button_2" at 1,354 size 78x58; TextOff 'Menu'
      on Release: ActivateScreen("Menu", 0)
   Button "Template_Button_3" at 401,354 size 78x58; TextOff 'Settings / Nastavania'
      on Release: ActivateScreen("Setting_DelayTime", 0)
   Button "Template_Button_4" at 481,354 size 78x58; TextOff 'Reset Faults Reset chýb'
      on Release: ResetBit("HMI_Control_ResetFaults")
      on Press: SetBit("HMI_Control_ResetFaults")
   Button "Template_Button_5" at 641,354 size 78x58; TextOff 'Text'; PictureOff "Graphic_7"
      on Release: function_a2a04561()
   Button "Template_Button_6" at 241,354 size 78x58; TextOff 'Status'
      on Release: ActivateScreen("StatusE", 0)
   Button "Alarms" at 161,354 size 78x58; TextOn 'Alarms / Alarmy'; TextOff 'Alarms / Alarmy'; PictureOn "AlarmDisplay_TP700_Comfort_TR"; PictureOff "AlarmDisplay_TP700_Comfort_TR"
      on Release: ActivateScreen("Alarm history_Enigma", 0)
   Button "Start screen" at 81,354 size 78x58; TextOn 'Start screen'; TextOff 'Start screen'; PictureOn "NavigateHome_TP700_Comfort_TR"; PictureOff "NavigateHome_TP700_Comfort_TR"
      on Release: ActivateScreen("MainScreen", 0)

Template "Template_Mirai" 800x414
   Button "Template_Button_1" at 561,354 size 78x58; TextOff 'System / Systém'
      on Release: ActivateScreen("SystemScreenM", 0)
   Button "Exit_1" at 721,354 size 78x58; TextOff 'Exit'; Authorization "User administration"; PictureOff "ExitRuntime_TP700_Comfort_TR"; PictureOn "ExitRuntime_TP700_Comfort_TR"
      on Release: StopRuntime(0)
   Button "Template_Button" at 321,354 size 78x58; TextOff 'Text'
   Button "Template_Button_9" at 1,354 size 78x58; TextOff 'Menu'
      on Release: ActivateScreen("Menu", 0)
   Button "Template_Button_10" at 401,354 size 78x58; TextOff 'Settings / Nastavania'
      on Release: ActivateScreen("SettingPrinter", 0)
   Button "Template_Button_11" at 481,354 size 78x58; TextOff 'Reset Faults Reset chýb'
      on Release: ResetBit("HMI_Control_ResetFaults")
      on Press: SetBit("HMI_Control_ResetFaults")
   Button "Template_Button_12" at 641,354 size 78x58; TextOff 'Text'; PictureOff "Graphic_7"
      on Release: function_a2a04561()
   Button "Template_Button_13" at 241,354 size 78x58; TextOff 'Status'
      on Release: ActivateScreen("StatusM", 0)
   Button "Alarms_1" at 161,354 size 78x58; TextOn 'Alarms / Alarmy'; TextOff 'Alarms / Alarmy'; PictureOn "AlarmDisplay_TP700_Comfort_TR"; PictureOff "AlarmDisplay_TP700_Comfort_TR"
      on Release: ActivateScreen("Alarm history_Mirai", 0)
   Button "Start screen_1" at 81,354 size 78x58; TextOn 'Start screen'; TextOff 'Start screen'; PictureOn "NavigateHome_TP700_Comfort_TR"; PictureOff "NavigateHome_TP700_Comfort_TR"
      on Release: ActivateScreen("Main", 0)

screen "Alarm history_Mirai" 800x414, template "Template_Mirai"
   on GenerateScreen: SetTag("screen_titles", 2)
   AlarmView "Alarm view_1" at 0,0 size 800x349

screen "SystemScreenM" 800x414, template "Template_Mirai"
   on GenerateScreen: SetTag("screen_titles", 20)
   Button "HmiScreenItemData_2" at 196,73 size 169x52; TextOn 'Projektinformationen / Project information / Informatii proiect / ข้อมูลโปรเจ็ค / Informácie o projekte'; TextOff 'Projektinformationen Project information Informatii proiect ข้อมูลโปรเจ็ค Informácie o projekte'; PictureOn "Navigates to Projektinformationen for HMI_1"; PictureOff "Graphic_1"
      on Press: ActivateScreen("ProjectInfo", 0)
   Button "HmiScreenItemData_3" at 435,201 size 169x52; TextOn 'Systemeinstellungen System settings Setarile de sistem Configurações de sistema ตั้งค่าระบบ Systémové nastavenia'; TextOff 'Systemeinstellungen System settings Setarile de sistem Configurações de sistema ตั้งค่าระบบ Systémové nastavenia'; Authorization "User administration"; PictureOff "Graphic_6"; PictureOn "Graphic_6"
      on Press: ActivateScreen("SystemSettings", 0)
   Button "HmiScreenItemData_4" at 196,137 size 169x52; TextOn 'Benutzerverwaltung User administration De administrare a utilizatorilor Administração de usuários การควบคุมผู้ใช้งาน Správa používateľov'; TextOff 'Benutzerverwaltung User administration De administrare a utilizatorilor Administração de usuários การควบคุมผู้ใช้งาน Správa používateľov'; Authorization "User administration"; PictureOff "Graphic_4"; PictureOn "Navigates to Benutzerverwaltung for HMI_1"
      on Press: ActivateScreen("UserAdmin", 0)
   Button "HmiScreenItemData_5" at 435,73 size 169x52; TextOn 'Systeminformationen / System information / Informatii sistem / Informação do sistema / ข้อมูลระบบ / Informácie o systéme'; TextOff 'Systeminformationen System information Informatii sistem Informação do sistema ข้อมูลระบบ Informácie o systéme'; PictureOn "Graphic_2"; PictureOff "Graphic_2"
      on Press: ActivateScreen("SystemInfo", 0)
   Button "HmiScreenItemData_6" at 435,137 size 169x52; TextOn 'Verschiedene Aufgaben Other tools Diverse activitati Various tasks งานอื่นๆ Iné nástroje'; TextOff 'Verschiedene Aufgaben Other tools Diverse activitati Various tasks งานอื่นๆ Iné nástroje'; PictureOn "Navigates to Verschiedene Aufgaben for HMI_1"; PictureOff "Graphic_5"
      on Press: ActivateScreen("OtherTools", 0)
   Button "HmiScreenItemData_1" at 195,201 size 169x52; TextOn 'Systemeinstellungen System diagnostics Setarile de sistem Configurações de sistema ตั้งค่าระบบ Diagnostika systému'; TextOff 'Systemeinstellungen System diagnostics Setarile de sistem Configurações de sistema ตั้งค่าระบบ Diagnostika systému'; PictureOff "Graphic_3"; PictureOn "Graphic_3"; Authorization "Operate"
      on Press: ActivateScreen("Diagnostic", 0)

screen "Setting_CameraM" 800x414, template "Template_Enigma"
   on GenerateScreen: SetTag("screen_titles", 54)
   IOField "I/O field_1" at 407,126 size 104x32; FormatPattern 9999
      ProcessValue <- "SP_HMI_Bag_Cam_Vertiacal_position"
   IOField "I/O field_2" at 407,202 size 104x32; FormatPattern s999
      ProcessValue <- "SP_HMI_Bag_Cam_Angle"
   IOField "I/O field_3" at 407,164 size 104x32; FormatPattern 9999
      ProcessValue <- "SP_HMI_Bag_Cam_Horizontal_position"
   TextField "Text field_1" at 299,126 size 104x32; Text 'A'
   TextField "Text field_2" at 299,164 size 104x32; Text 'B'
   TextField "Text field_3" at 299,202 size 104x32; Text 'C'
   TextField "Text field_4" at 623,126 size 36x32; Text 'mm'
   TextField "Text field_5" at 623,164 size 36x32; Text 'mm'
   TextField "Text field_6" at 623,202 size 36x32; Text '°'
   TextField "Text field_18" at 419,90 size 80x32; Text 'BAG / SÁČOK'
   TextField "Text field_19" at 523,90 size 80x32; Text 'BOX / KRABICA'
   IOField "I/O field_8" at 515,126 size 104x32; FormatPattern 9999
      ProcessValue <- "SP_HMI_Box_Cam_Vertiacal_position"
   IOField "I/O field_9" at 515,202 size 104x32; FormatPattern s999
      ProcessValue <- "SP_HMI_Box_Cam_Angle"
   IOField "I/O field_10" at 515,164 size 104x32; FormatPattern 9999
      ProcessValue <- "SP_HMI_Box_Cam_Horizontal_position"
   Button "Button_7" at 8,313 size 152x32; TextOff 'Back / Späť'
      on Click: ActivateScreen("Setting_DelayTimeM", 0)
   GraphicView "Graphic view_1" at 20,53 size 224x212; Picture "CognexDatamanEdited_3"
   TextField "Text field_10" at 18,144 size 32x40; Text 'A'
   TextField "Text field_11" at 102,31 size 32x40; Text 'B'
   TextField "Text field_12" at 179,38 size 32x40; Text 'C'
   TextField "Text field_7" at 288,8 size 376x62; Text 'Camera position: / Pozícia kamery: / 配方名'
   GraphicIOField "Graphic I/O field_1" at 408,243 size 32x32; PictureList "On_Off_NonEditable"
      ProcessValue <- "SP_HMI_Enigma_off"
   TextField "Text field_14" at 299,243 size 104x32; Text 'Enigma'
   GraphicIOField "Graphic I/O field_2" at 624,243 size 32x32; PictureList "On_Off_NonEditable"
      ProcessValue <- "SP_HMI_Mirai_off"
   TextField "Text field_20" at 515,243 size 104x32; Text 'Mirai'

PopupScreen "AutoSelectRecipeFailed" 800x480
   TextField "Text field_2" at 200,128 size 400x80; Text 'Automatické načítavanie receptu zlyhalo. Zvoľte a nahrajte recept manuálne alebo požadovaný recept vytvorte! Auto recipe loading failed. Select and load recipe manually or create a required recipe.'
   Button "Button_3" at 362,216 size 76x32; TextOff 'OK'
      on Click: function_efd93a16("AutoSelectRecipeFailed", 0, 0, 0, -1, 1)

VB script "Rec_EmergencyReset"
   SmartTags("Rec_DeleteResult") = 0
   SmartTags("Rec_EditResult") = 0
   SmartTags("Rec_AutoSelectResult") = 0
   'SmartTags("Rec_ExportResult") = 0
   'SmartTags("Rec_ImportResult") = 0
   SmartTags("Rec_LoadResult") = 0
   SmartTags("Rec_ReadSPResult") = 0
   SmartTags("Rec_SaveResult") = 0
   SmartTags("Rec_ViewResult") = 0
   SmartTags("Rec_FunctionUsed") = 0

VB script "Rec_SafeDelete"
   If SmartTags("Rec_SelectedRecipe") <> "" Then
   	cbbc2fc1-4696-421a-97b4-46a748b4d57f 1, SmartTags("Rec_SelectedRecipe"), $3$hmiOn$, $3$hmiOn$, Rec_DeleteResult
   Else
   	SmartTags("Rec_DeleteResult") = -1
   End If

VB script "Rec_SafeEdit"
   If SmartTags("Rec_SelectedRecipe") <> "" Then
   	b431313b-d6b5-4a28-b630-23a386ef7180 1, SmartTags("Rec_SelectedRecipe"), Rec_EditResult
   Else
   	SmartTags("Rec_EditResult") = -1
   End If

VB script "Rec_SafeLoad"
   If SmartTags("Rec_SelectedRecipe") <> "" Then
   	eba64363-2936-407c-9a7c-00964fb48e05 1, SmartTags("Rec_SelectedRecipe"), $3$hmiOn$, Rec_LoadResult
   Else
   	SmartTags("Rec_LoadResult") = -1
   End If

VB script "Rec_SafeSave"
   If SmartTags("Rec_SelectedRecipe") <> "" Then
   	f38ba6b2-0c13-4a6f-acab-73f2fde9baea 1, SmartTags("Rec_SelectedRecipe"), $3$hmiOverwriteWithConfirmation$, $3$hmiOn$, Rec_SaveResult
   Else
   	SmartTags("Rec_SaveResult") = -1
   End If

VB script "Rec_SafeView"
   If SmartTags("Rec_SelectedRecipe") <> "" Then
   	b431313b-d6b5-4a28-b630-23a386ef7180 1, SmartTags("Rec_SelectedRecipe"), Rec_ViewResult
   Else
   	SmartTags("Rec_ViewResult") = -1
   End If

VB script "AutoLoginOperator"
   If (SmartTags("liuser") = "") Or (SmartTags("initDone") = 0) Then
   	a9b89908-c625-4370-ad53-4ebfb8d097d7 autoPwd, autoUser
   	SmartTags("autoPwd") = "operator"
   	SmartTags("autoUser") = "operator"
   	SmartTags("initDone") = 1
   End If

VB script "Rec_AutoSelectRecipe"
   	If SmartTags("FindRecipe") Then
   		b21d3eaf-4e31-425c-ad1a-ba4e4002cacc Rec_FunctionUsed, 3
   		
   		eba64363-2936-407c-9a7c-00964fb48e05 1, SmartTags("PlainHandle_DB_NewArticleNum"), $3$hmiOn$, Rec_AutoSelectResult
   		
   		While SmartTags("Rec_AutoSelectResult") = 2
   				' Wait to operation complete.
   		Wend
   		
   		If SmartTags ("Rec_AutoSelectResult") = 4 Then
   			bfde4b54-0db7-4817-8032-87127bf19bb9 "Nový recept bol automaticky nahratý do PLC."
   			db265680-6104-4a2a-bb94-41ffdc16be82 HMI_Control_NewRecipeLoaded			
   		Else
   			bfde4b54-0db7-4817-8032-87127bf19bb9 "Pri automatickom nahrávaní receptu nastala chyba."
   			efd93a16-2665-4b85-bcb9-25eddcb7b6f4  AutoSelectRecipeFailed, 0, 0, $3$hmiOn$, $3$hmiAnimationOff$, $3$hmiMedium$
   			db265680-6104-4a2a-bb94-41ffdc16be82 HMI_Control_AutoRecipeFailed
   		End If
   		
   		SmartTags("Rec_AutoSelectResult") = 0
   	End If

scheduled task "UserChange"
   on Action: function_f41c6f6c("liuser"); "AutoLoginOperator"()
*)